REGION Network 25: RESET TEMPO DE OPERAÇÃO (HORAS)
   RUNG wire#powerrail
      Contact( #AUX09 )
      wire#w1
      { S7_GenerateENO := "TRUE" } Move(in := 0, out1 => #HOR)
   END_RUNG
   RUNG wire#powerrail
      Contact( #CRTO )
   END_RUNG wire#w1
   // the same network as SCL:
   IF #AUX09 OR #CRTO THEN #HOR := 0; END_IF;
END_REGION

REGION Network 26 (STL): ESCRITA DOS DADOS NO INVERSOR (PALAVRA DE COMANDO)
         A     "AlwaysTRUE";
         =     #CTW.DCbrakeRamp;
         =     #CTW.Coasting;
         =     #CTW.Enable_Ramp;
         =     #CTW.Enable_ramp_generator;
         =     #CTW.Control_plc;  //Valida setpoint


         A     #CL;
         =     #CTW.Start;  //LIGA/DESL

         A     #CL;
         A     #AUX10;
         A     #HAR;
         =     #CTW.Start_reverse;  //LIGA/DESL REVERSO


         A     #RESET;
         AN    #CL;
         =     #CTW.Reset;  //RESET
END_REGION
END_FUNCTION_BLOCK

FUNCTION_BLOCK "PDIR"   // FB207, LAD
{ S7_Optimized_Access := 'FALSE' }
VERSION : 0.1
   VAR_INPUT
      ML : Bool;
      MR : Bool;
      DL : Bool;
      MF1 : Bool;
      MF2 : Bool;
      HM : Bool;
      HA : Bool;
      CMA : Bool;
      CLM : Bool;
      CDM : Bool;
      CRF : Bool;
      CRTO : Bool;
      CL1S : Bool;
   END_VAR
   VAR_OUTPUT
      YFPP : Bool;
      YF : Bool;
      CL : Bool;
   END_VAR
   VAR_IN_OUT
      SEG : Int;
      MIN : Int;
      HOR : Int;
   END_VAR
   VAR
      AUX01 : Bool;
      AUX02 : Bool;
      AUX03 : Bool;
      AUX04 : Bool;
      AUX05 : Bool;
      AUX06 : Bool;
      AUX07 : Bool;
      AUX08 : Bool;
      AUX09 : Bool;
      P60S : Bool;
      P60M : Bool;
      PFHO : Bool;
      TPP1 : TON_TIME;
      TPP2 : TON_TIME;
   END_VAR
   VAR_TEMP
      TEMP0 : Bool;
      TEMP1 : Bool;
      ET_TPP1 : Time;
      ET_TPP2 : Time;
   END_VAR
   VAR_TEMP   // added for the SCL form of the ladder/FBD networks
      _w1 : Bool;
      _w2 : Bool;
      _w3 : Bool;
      _w4 : Bool;
   END_VAR
BEGIN

REGION Network 1: Falha na partida
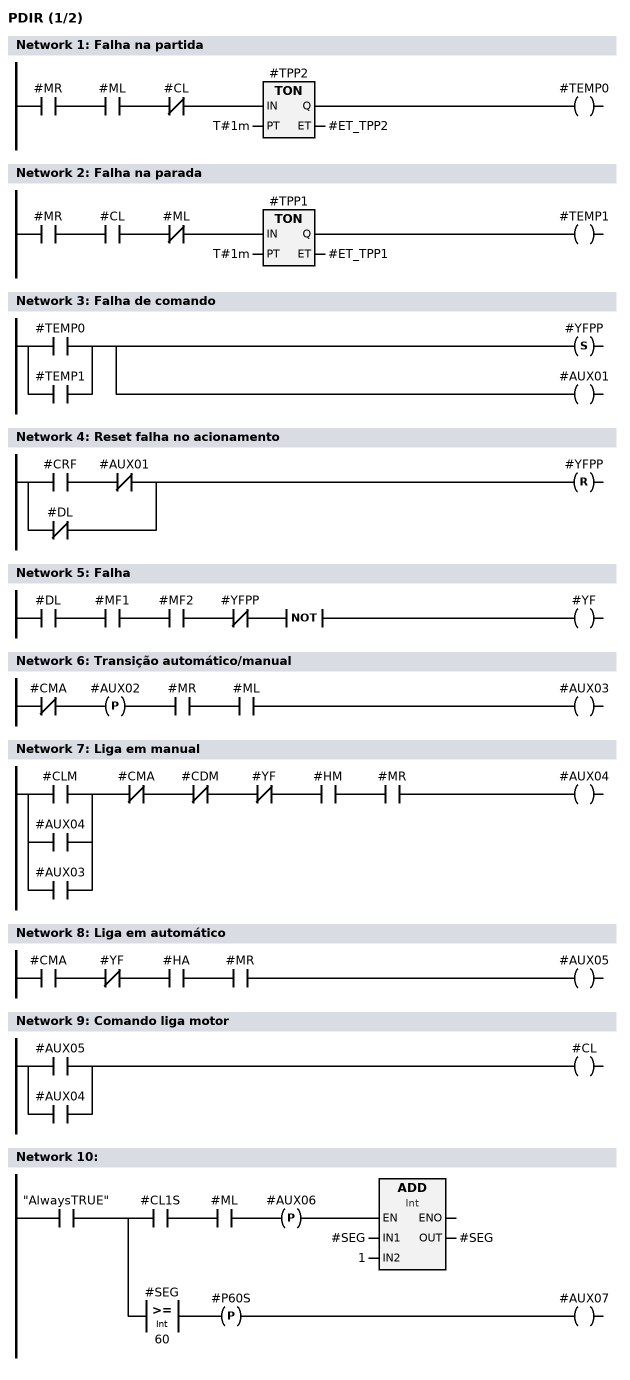
   #TPP2(IN := #MR AND #ML AND NOT #CL, PT := T#1m, ET => #ET_TPP2);   // TON
   #TEMP0 := #TPP2.Q;
END_REGION

REGION Network 2: Falha na parada
   #TPP1(IN := #MR AND #CL AND NOT #ML, PT := T#1m, ET => #ET_TPP1);   // TON
   #TEMP1 := #TPP1.Q;
END_REGION

REGION Network 3: Falha de comando
   RUNG wire#powerrail
      Contact( #TEMP0 )
      wire#w1
      S_Coil( #YFPP )
   END_RUNG
   RUNG wire#powerrail
      Contact( #TEMP1 )
   END_RUNG wire#w1
   RUNG wire#w1
      Coil( #AUX01 )
   END_RUNG
   // the same network as SCL:
   #_w1 := #TEMP0 OR #TEMP1;
   IF #_w1 THEN #YFPP := TRUE; END_IF;
   #AUX01 := #_w1;
END_REGION

REGION Network 4: Reset falha no acionamento
   RUNG wire#powerrail
      Contact( #CRF )
      I_Contact( #AUX01 )
      wire#w1
      R_Coil( #YFPP )
   END_RUNG
   RUNG wire#powerrail
      I_Contact( #DL )
   END_RUNG wire#w1
   // the same network as SCL:
   IF (#CRF AND NOT #AUX01) OR NOT #DL THEN #YFPP := FALSE; END_IF;
END_REGION

REGION Network 5: Falha
   RUNG wire#powerrail
      Contact( #DL )
      Contact( #MF1 )
      Contact( #MF2 )
      I_Contact( #YFPP )
      Not()
      Coil( #YF )
   END_RUNG
   // the same network as SCL:
   #YF := NOT (#DL AND #MF1 AND #MF2 AND NOT #YFPP);
END_REGION

REGION Network 6: Transição automático/manual
   RUNG wire#powerrail
      I_Contact( #CMA )
      P_Trig( #AUX02 )
      Contact( #MR )
      Contact( #ML )
      Coil( #AUX03 )
   END_RUNG
   // the same network as SCL:
   #_w1 := NOT #CMA AND NOT #AUX02;   // rising edge
   #AUX02 := NOT #CMA;
   #AUX03 := #_w1 AND #MR AND #ML;
END_REGION

REGION Network 7: Liga em manual
   RUNG wire#powerrail
      Contact( #CLM )
      wire#w1
      I_Contact( #CMA )
      I_Contact( #CDM )
      I_Contact( #YF )
      Contact( #HM )
      Contact( #MR )
      Coil( #AUX04 )
   END_RUNG
   RUNG wire#powerrail
      Contact( #AUX04 )
   END_RUNG wire#w1
   RUNG wire#powerrail
      Contact( #AUX03 )
   END_RUNG wire#w1
   // the same network as SCL:
   #AUX04 := (#CLM OR #AUX04 OR #AUX03) AND NOT #CMA AND NOT #CDM AND NOT #YF AND #HM AND #MR;
END_REGION

REGION Network 8: Liga em automático
   RUNG wire#powerrail
      Contact( #CMA )
      I_Contact( #YF )
      Contact( #HA )
      Contact( #MR )
      Coil( #AUX05 )
   END_RUNG
   // the same network as SCL:
   #AUX05 := #CMA AND NOT #YF AND #HA AND #MR;
END_REGION

REGION Network 9: Comando liga motor
   RUNG wire#powerrail
      Contact( #AUX05 )
      wire#w1
      Coil( #CL )
   END_RUNG
   RUNG wire#powerrail
      Contact( #AUX04 )
   END_RUNG wire#w1
   // the same network as SCL:
   #CL := #AUX05 OR #AUX04;
END_REGION

REGION Network 10
   RUNG wire#powerrail
      Contact( "AlwaysTRUE" )
      wire#w1
      Contact( #CL1S )
      Contact( #ML )
      P_Trig( #AUX06 )
      { S7_Templates := "SrcType := Int"; S7_GenerateENO := "TRUE" } Add(in1 := #SEG, in2 := 1, out => #SEG)
   END_RUNG
   RUNG wire#w1
      { S7_Templates := "SrcType := Int" } GE_Contact(in1 := #SEG, in2 := 60)
      P_Trig( #P60S )
      Coil( #AUX07 )
   END_RUNG
   // the same network as SCL:
   #_w1 := "AlwaysTRUE" AND #CL1S AND #ML;
   #_w2 := #_w1 AND NOT #AUX06;   // rising edge
   #AUX06 := #_w1;
   IF #_w2 THEN #SEG := #SEG + 1; END_IF;
   #_w3 := "AlwaysTRUE" AND (#SEG >= 60);
   #_w4 := #_w3 AND NOT #P60S;   // rising edge
   #P60S := #_w3;
   #AUX07 := #_w4;
END_REGION

REGION Network 11
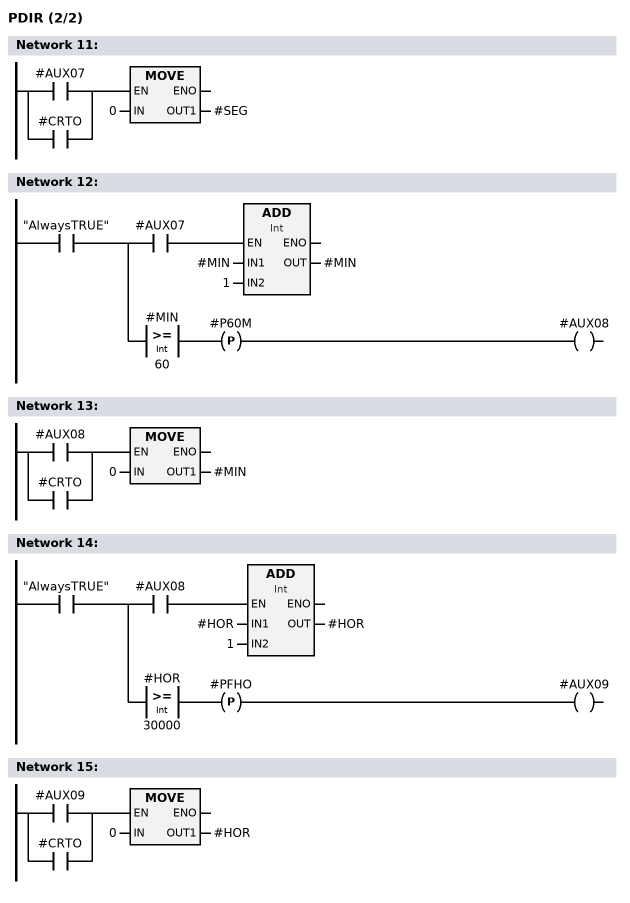
   RUNG wire#powerrail
      Contact( #AUX07 )
      wire#w1
      { S7_GenerateENO := "TRUE" } Move(in := 0, out1 => #SEG)
   END_RUNG
   RUNG wire#powerrail
      Contact( #CRTO )
   END_RUNG wire#w1
   // the same network as SCL:
   IF #AUX07 OR #CRTO THEN #SEG := 0; END_IF;
END_REGION

REGION Network 12
   RUNG wire#powerrail
      Contact( "AlwaysTRUE" )
      wire#w1
      Contact( #AUX07 )
      { S7_Templates := "SrcType := Int"; S7_GenerateENO := "TRUE" } Add(in1 := #MIN, in2 := 1, out => #MIN)
   END_RUNG
   RUNG wire#w1
      { S7_Templates := "SrcType := Int" } GE_Contact(in1 := #MIN, in2 := 60)
      P_Trig( #P60M )
      Coil( #AUX08 )
   END_RUNG
   // the same network as SCL:
   IF "AlwaysTRUE" AND #AUX07 THEN #MIN := #MIN + 1; END_IF;
   #_w1 := "AlwaysTRUE" AND (#MIN >= 60);
   #_w2 := #_w1 AND NOT #P60M;   // rising edge
   #P60M := #_w1;
   #AUX08 := #_w2;
END_REGION

REGION Network 13
   RUNG wire#powerrail
      Contact( #AUX08 )
      wire#w1
      { S7_GenerateENO := "TRUE" } Move(in := 0, out1 => #MIN)
   END_RUNG
   RUNG wire#powerrail
      Contact( #CRTO )
   END_RUNG wire#w1
   // the same network as SCL:
   IF #AUX08 OR #CRTO THEN #MIN := 0; END_IF;
END_REGION

REGION Network 14
   RUNG wire#powerrail
      Contact( "AlwaysTRUE" )
      wire#w1
      Contact( #AUX08 )
      { S7_Templates := "SrcType := Int"; S7_GenerateENO := "TRUE" } Add(in1 := #HOR, in2 := 1, out => #HOR)
   END_RUNG
   RUNG wire#w1
      { S7_Templates := "SrcType := Int" } GE_Contact(in1 := #HOR, in2 := 30000)
      P_Trig( #PFHO )
      Coil( #AUX09 )
   END_RUNG
   // the same network as SCL:
   IF "AlwaysTRUE" AND #AUX08 THEN #HOR := #HOR + 1; END_IF;
   #_w1 := "AlwaysTRUE" AND (#HOR >= 30000);
   #_w2 := #_w1 AND NOT #PFHO;   // rising edge
   #PFHO := #_w1;
   #AUX09 := #_w2;
END_REGION

REGION Network 15
   RUNG wire#powerrail
      Contact( #AUX09 )
      wire#w1
      { S7_GenerateENO := "TRUE" } Move(in := 0, out1 => #HOR)
   END_RUNG
   RUNG wire#powerrail
      Contact( #CRTO )
   END_RUNG wire#w1
   // the same network as SCL:
   IF #AUX09 OR #CRTO THEN #HOR := 0; END_IF;
END_REGION
END_FUNCTION_BLOCK

FUNCTION "IO" : Void   // FC1, LAD
{ S7_Optimized_Access := 'TRUE' }
VERSION : 0.1
BEGIN

REGION Network 1: Status e alarme elevatória principal 1
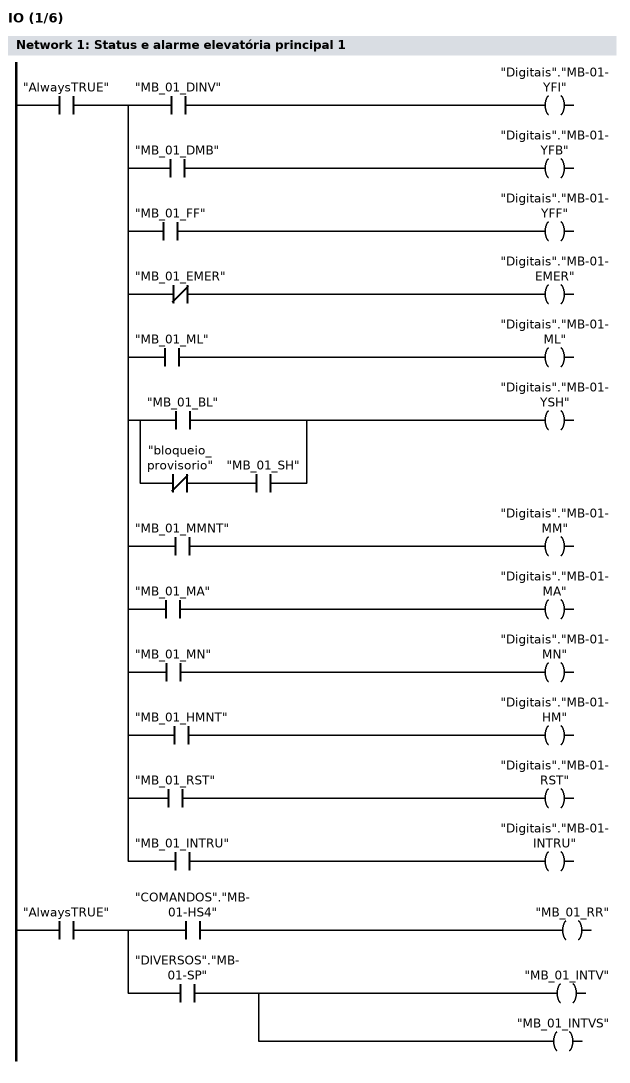
   RUNG wire#powerrail
      Contact( "AlwaysTRUE" )
      wire#w1
      Contact( "MB_01_DINV" )
      Coil( "Digitais"."MB-01-YFI" )
   END_RUNG
   RUNG wire#w1
      Contact( "MB_01_DMB" )
      Coil( "Digitais"."MB-01-YFB" )
   END_RUNG
   RUNG wire#w1
      Contact( "MB_01_FF" )
      Coil( "Digitais"."MB-01-YFF" )
   END_RUNG
   RUNG wire#w1
      I_Contact( "MB_01_EMER" )
      Coil( "Digitais"."MB-01-EMER" )
   END_RUNG
   RUNG wire#w1
      Contact( "MB_01_ML" )
      Coil( "Digitais"."MB-01-ML" )
   END_RUNG
   RUNG wire#w1
      Contact( "MB_01_BL" )
      wire#w2
      Coil( "Digitais"."MB-01-YSH" )
   END_RUNG
   RUNG wire#w1
      I_Contact( "bloqueio_provisorio" )
      Contact( "MB_01_SH" )
   END_RUNG wire#w2
   RUNG wire#w1
      Contact( "MB_01_MMNT" )
      Coil( "Digitais"."MB-01-MM" )
   END_RUNG
   RUNG wire#w1
      Contact( "MB_01_MA" )
      Coil( "Digitais"."MB-01-MA" )
   END_RUNG
   RUNG wire#w1
      Contact( "MB_01_MN" )
      Coil( "Digitais"."MB-01-MN" )
   END_RUNG
   RUNG wire#w1
      Contact( "MB_01_HMNT" )
      Coil( "Digitais"."MB-01-HM" )
   END_RUNG
   RUNG wire#w1
      Contact( "MB_01_RST" )
      Coil( "Digitais"."MB-01-RST" )
   END_RUNG
   RUNG wire#w1
      Contact( "MB_01_INTRU" )
      Coil( "Digitais"."MB-01-INTRU" )
   END_RUNG
   RUNG wire#powerrail
      Contact( "AlwaysTRUE" )
      wire#w3
      Contact( "COMANDOS"."MB-01-HS4" )
      Coil( "MB_01_RR" )
   END_RUNG
   RUNG wire#w3
      Contact( "DIVERSOS"."MB-01-SP" )
      wire#w4
      Coil( "MB_01_INTV" )
   END_RUNG
   RUNG wire#w4
      Coil( "MB_01_INTVS" )
   END_RUNG
   // the same network as SCL:
   "Digitais"."MB-01-YFI" := "AlwaysTRUE" AND "MB_01_DINV";
   "Digitais"."MB-01-YFB" := "AlwaysTRUE" AND "MB_01_DMB";
   "Digitais"."MB-01-YFF" := "AlwaysTRUE" AND "MB_01_FF";
   "Digitais"."MB-01-EMER" := "AlwaysTRUE" AND NOT "MB_01_EMER";
   "Digitais"."MB-01-ML" := "AlwaysTRUE" AND "MB_01_ML";
   "Digitais"."MB-01-YSH" := "AlwaysTRUE" AND ("MB_01_BL" OR (NOT "bloqueio_provisorio" AND "MB_01_SH"));
   "Digitais"."MB-01-MM" := "AlwaysTRUE" AND "MB_01_MMNT";
   "Digitais"."MB-01-MA" := "AlwaysTRUE" AND "MB_01_MA";
   "Digitais"."MB-01-MN" := "AlwaysTRUE" AND "MB_01_MN";
   "Digitais"."MB-01-HM" := "AlwaysTRUE" AND "MB_01_HMNT";
   "Digitais"."MB-01-RST" := "AlwaysTRUE" AND "MB_01_RST";
   "Digitais"."MB-01-INTRU" := "AlwaysTRUE" AND "MB_01_INTRU";
   "MB_01_RR" := "AlwaysTRUE" AND "COMANDOS"."MB-01-HS4";
   "MB_01_INTV" := "AlwaysTRUE" AND "DIVERSOS"."MB-01-SP";
   "MB_01_INTVS" := "MB_01_INTV";
END_REGION

REGION Network 2: Status e alarme elevatória principal 2
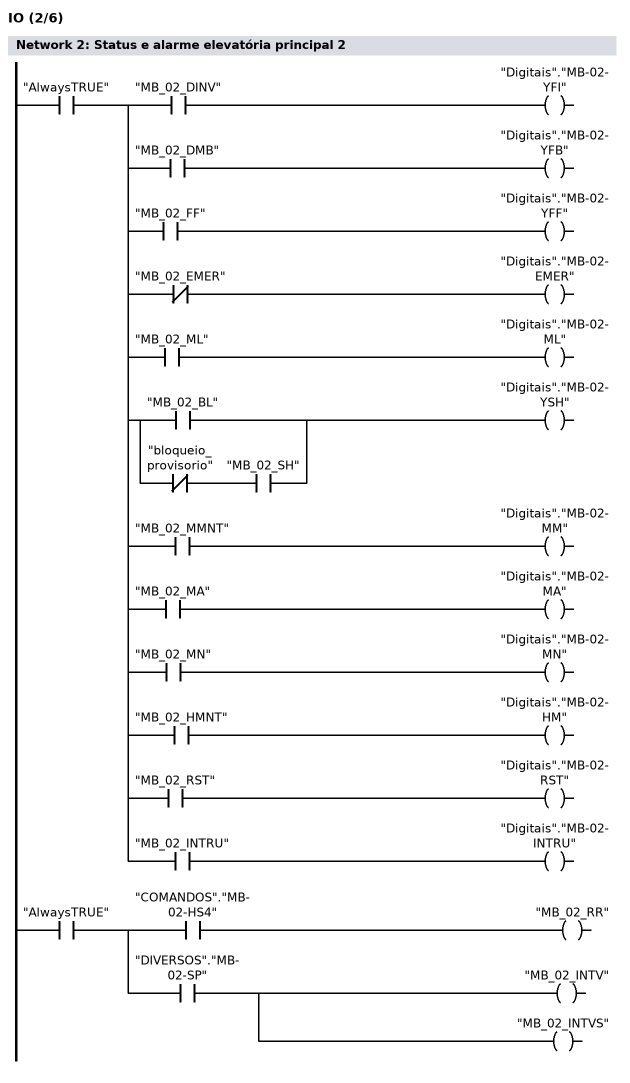
   RUNG wire#powerrail
      Contact( "AlwaysTRUE" )
      wire#w1
      Contact( "MB_02_DINV" )
      Coil( "Digitais"."MB-02-YFI" )
   END_RUNG
   RUNG wire#w1
      Contact( "MB_02_DMB" )
      Coil( "Digitais"."MB-02-YFB" )
   END_RUNG
   RUNG wire#w1
      Contact( "MB_02_FF" )
      Coil( "Digitais"."MB-02-YFF" )
   END_RUNG
   RUNG wire#w1
      I_Contact( "MB_02_EMER" )
      Coil( "Digitais"."MB-02-EMER" )
   END_RUNG
   RUNG wire#w1
      Contact( "MB_02_ML" )
      Coil( "Digitais"."MB-02-ML" )
   END_RUNG
   RUNG wire#w1
      Contact( "MB_02_BL" )
      wire#w2
      Coil( "Digitais"."MB-02-YSH" )
   END_RUNG
   RUNG wire#w1
      I_Contact( "bloqueio_provisorio" )
      Contact( "MB_02_SH" )
   END_RUNG wire#w2
   RUNG wire#w1
      Contact( "MB_02_MMNT" )
      Coil( "Digitais"."MB-02-MM" )
   END_RUNG
   RUNG wire#w1
      Contact( "MB_02_MA" )
      Coil( "Digitais"."MB-02-MA" )
   END_RUNG
   RUNG wire#w1
      Contact( "MB_02_MN" )
      Coil( "Digitais"."MB-02-MN" )
   END_RUNG
   RUNG wire#w1
      Contact( "MB_02_HMNT" )
      Coil( "Digitais"."MB-02-HM" )
   END_RUNG
   RUNG wire#w1
      Contact( "MB_02_RST" )
      Coil( "Digitais"."MB-02-RST" )
   END_RUNG
   RUNG wire#w1
      Contact( "MB_02_INTRU" )
      Coil( "Digitais"."MB-02-INTRU" )
   END_RUNG
   RUNG wire#powerrail
      Contact( "AlwaysTRUE" )
      wire#w3
      Contact( "COMANDOS"."MB-02-HS4" )
      Coil( "MB_02_RR" )
   END_RUNG
   RUNG wire#w3
      Contact( "DIVERSOS"."MB-02-SP" )
      wire#w4
      Coil( "MB_02_INTV" )
   END_RUNG
   RUNG wire#w4
      Coil( "MB_02_INTVS" )
   END_RUNG
   // the same network as SCL:
   "Digitais"."MB-02-YFI" := "AlwaysTRUE" AND "MB_02_DINV";
   "Digitais"."MB-02-YFB" := "AlwaysTRUE" AND "MB_02_DMB";
   "Digitais"."MB-02-YFF" := "AlwaysTRUE" AND "MB_02_FF";
   "Digitais"."MB-02-EMER" := "AlwaysTRUE" AND NOT "MB_02_EMER";
   "Digitais"."MB-02-ML" := "AlwaysTRUE" AND "MB_02_ML";
   "Digitais"."MB-02-YSH" := "AlwaysTRUE" AND ("MB_02_BL" OR (NOT "bloqueio_provisorio" AND "MB_02_SH"));
   "Digitais"."MB-02-MM" := "AlwaysTRUE" AND "MB_02_MMNT";
   "Digitais"."MB-02-MA" := "AlwaysTRUE" AND "MB_02_MA";
   "Digitais"."MB-02-MN" := "AlwaysTRUE" AND "MB_02_MN";
   "Digitais"."MB-02-HM" := "AlwaysTRUE" AND "MB_02_HMNT";
   "Digitais"."MB-02-RST" := "AlwaysTRUE" AND "MB_02_RST";
   "Digitais"."MB-02-INTRU" := "AlwaysTRUE" AND "MB_02_INTRU";
   "MB_02_RR" := "AlwaysTRUE" AND "COMANDOS"."MB-02-HS4";
   "MB_02_INTV" := "AlwaysTRUE" AND "DIVERSOS"."MB-02-SP";
   "MB_02_INTVS" := "MB_02_INTV";
END_REGION

REGION Network 3: Status e alarme elevatória principal 3
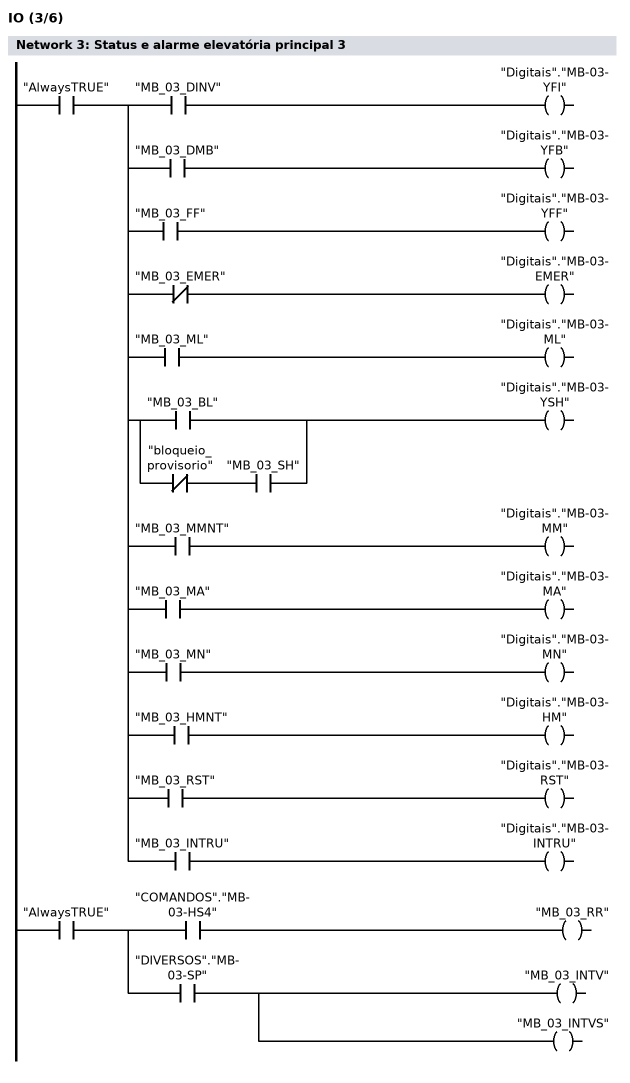
   RUNG wire#powerrail
      Contact( "AlwaysTRUE" )
      wire#w1
      Contact( "MB_03_DINV" )
      Coil( "Digitais"."MB-03-YFI" )
   END_RUNG
   RUNG wire#w1
      Contact( "MB_03_DMB" )
      Coil( "Digitais"."MB-03-YFB" )
   END_RUNG
   RUNG wire#w1
      Contact( "MB_03_FF" )
      Coil( "Digitais"."MB-03-YFF" )
   END_RUNG
   RUNG wire#w1
      I_Contact( "MB_03_EMER" )
      Coil( "Digitais"."MB-03-EMER" )
   END_RUNG
   RUNG wire#w1
      Contact( "MB_03_ML" )
      Coil( "Digitais"."MB-03-ML" )
   END_RUNG
   RUNG wire#w1
      Contact( "MB_03_BL" )
      wire#w2
      Coil( "Digitais"."MB-03-YSH" )
   END_RUNG
   RUNG wire#w1
      I_Contact( "bloqueio_provisorio" )
      Contact( "MB_03_SH" )
   END_RUNG wire#w2
   RUNG wire#w1
      Contact( "MB_03_MMNT" )
      Coil( "Digitais"."MB-03-MM" )
   END_RUNG
   RUNG wire#w1
      Contact( "MB_03_MA" )
      Coil( "Digitais"."MB-03-MA" )
   END_RUNG
   RUNG wire#w1
      Contact( "MB_03_MN" )
      Coil( "Digitais"."MB-03-MN" )
   END_RUNG
   RUNG wire#w1
      Contact( "MB_03_HMNT" )
      Coil( "Digitais"."MB-03-HM" )
   END_RUNG
   RUNG wire#w1
      Contact( "MB_03_RST" )
      Coil( "Digitais"."MB-03-RST" )
   END_RUNG
   RUNG wire#w1
      Contact( "MB_03_INTRU" )
      Coil( "Digitais"."MB-03-INTRU" )
   END_RUNG
   RUNG wire#powerrail
      Contact( "AlwaysTRUE" )
      wire#w3
      Contact( "COMANDOS"."MB-03-HS4" )
      Coil( "MB_03_RR" )
   END_RUNG
   RUNG wire#w3
      Contact( "DIVERSOS"."MB-03-SP" )
      wire#w4
      Coil( "MB_03_INTV" )
   END_RUNG
   RUNG wire#w4
      Coil( "MB_03_INTVS" )
   END_RUNG
   // the same network as SCL:
   "Digitais"."MB-03-YFI" := "AlwaysTRUE" AND "MB_03_DINV";
   "Digitais"."MB-03-YFB" := "AlwaysTRUE" AND "MB_03_DMB";
   "Digitais"."MB-03-YFF" := "AlwaysTRUE" AND "MB_03_FF";
   "Digitais"."MB-03-EMER" := "AlwaysTRUE" AND NOT "MB_03_EMER";
   "Digitais"."MB-03-ML" := "AlwaysTRUE" AND "MB_03_ML";
   "Digitais"."MB-03-YSH" := "AlwaysTRUE" AND ("MB_03_BL" OR (NOT "bloqueio_provisorio" AND "MB_03_SH"));
   "Digitais"."MB-03-MM" := "AlwaysTRUE" AND "MB_03_MMNT";
   "Digitais"."MB-03-MA" := "AlwaysTRUE" AND "MB_03_MA";
   "Digitais"."MB-03-MN" := "AlwaysTRUE" AND "MB_03_MN";
   "Digitais"."MB-03-HM" := "AlwaysTRUE" AND "MB_03_HMNT";
   "Digitais"."MB-03-RST" := "AlwaysTRUE" AND "MB_03_RST";
   "Digitais"."MB-03-INTRU" := "AlwaysTRUE" AND "MB_03_INTRU";
   "MB_03_RR" := "AlwaysTRUE" AND "COMANDOS"."MB-03-HS4";
   "MB_03_INTV" := "AlwaysTRUE" AND "DIVERSOS"."MB-03-SP";
   "MB_03_INTVS" := "MB_03_INTV";
END_REGION

REGION Network 4: Status e alarme elevatória principal 4
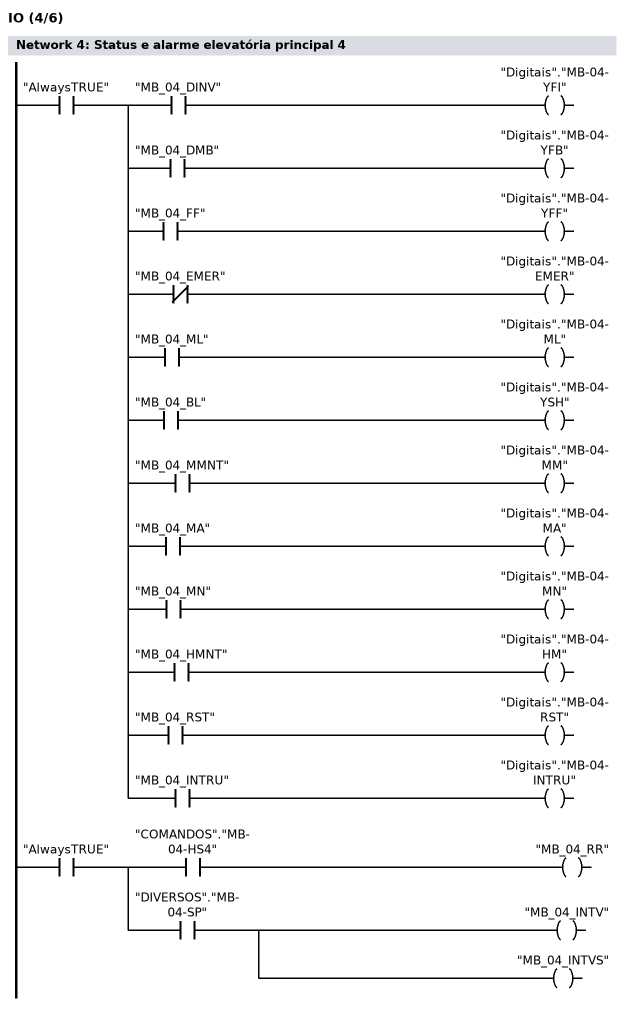
   RUNG wire#powerrail
      Contact( "AlwaysTRUE" )
      wire#w1
      Contact( "MB_04_DINV" )
      Coil( "Digitais"."MB-04-YFI" )
   END_RUNG
   RUNG wire#w1
      Contact( "MB_04_DMB" )
      Coil( "Digitais"."MB-04-YFB" )
   END_RUNG
   RUNG wire#w1
      Contact( "MB_04_FF" )
      Coil( "Digitais"."MB-04-YFF" )
   END_RUNG
   RUNG wire#w1
      I_Contact( "MB_04_EMER" )
      Coil( "Digitais"."MB-04-EMER" )
   END_RUNG
   RUNG wire#w1
      Contact( "MB_04_ML" )
      Coil( "Digitais"."MB-04-ML" )
   END_RUNG
   RUNG wire#w1
      Contact( "MB_04_BL" )
      Coil( "Digitais"."MB-04-YSH" )
   END_RUNG
   RUNG wire#w1
      Contact( "MB_04_MMNT" )
      Coil( "Digitais"."MB-04-MM" )
   END_RUNG
   RUNG wire#w1
      Contact( "MB_04_MA" )
      Coil( "Digitais"."MB-04-MA" )
   END_RUNG
   RUNG wire#w1
      Contact( "MB_04_MN" )
      Coil( "Digitais"."MB-04-MN" )
   END_RUNG
   RUNG wire#w1
      Contact( "MB_04_HMNT" )
      Coil( "Digitais"."MB-04-HM" )
   END_RUNG
   RUNG wire#w1
      Contact( "MB_04_RST" )
      Coil( "Digitais"."MB-04-RST" )
   END_RUNG
   RUNG wire#w1
      Contact( "MB_04_INTRU" )
      Coil( "Digitais"."MB-04-INTRU" )
   END_RUNG
   RUNG wire#powerrail
      Contact( "AlwaysTRUE" )
      wire#w2
      Contact( "COMANDOS"."MB-04-HS4" )
      Coil( "MB_04_RR" )
   END_RUNG
   RUNG wire#w2
      Contact( "DIVERSOS"."MB-04-SP" )
      wire#w3
      Coil( "MB_04_INTV" )
   END_RUNG
   RUNG wire#w3
      Coil( "MB_04_INTVS" )
   END_RUNG
   // the same network as SCL:
   "Digitais"."MB-04-YFI" := "AlwaysTRUE" AND "MB_04_DINV";
   "Digitais"."MB-04-YFB" := "AlwaysTRUE" AND "MB_04_DMB";
   "Digitais"."MB-04-YFF" := "AlwaysTRUE" AND "MB_04_FF";
   "Digitais"."MB-04-EMER" := "AlwaysTRUE" AND NOT "MB_04_EMER";
   "Digitais"."MB-04-ML" := "AlwaysTRUE" AND "MB_04_ML";
   "Digitais"."MB-04-YSH" := "AlwaysTRUE" AND "MB_04_BL";
   "Digitais"."MB-04-MM" := "AlwaysTRUE" AND "MB_04_MMNT";
   "Digitais"."MB-04-MA" := "AlwaysTRUE" AND "MB_04_MA";
   "Digitais"."MB-04-MN" := "AlwaysTRUE" AND "MB_04_MN";
   "Digitais"."MB-04-HM" := "AlwaysTRUE" AND "MB_04_HMNT";
   "Digitais"."MB-04-RST" := "AlwaysTRUE" AND "MB_04_RST";
   "Digitais"."MB-04-INTRU" := "AlwaysTRUE" AND "MB_04_INTRU";
   "MB_04_RR" := "AlwaysTRUE" AND "COMANDOS"."MB-04-HS4";
   "MB_04_INTV" := "AlwaysTRUE" AND "DIVERSOS"."MB-04-SP";
   "MB_04_INTVS" := "MB_04_INTV";
END_REGION

REGION Network 5: Status e alarme PCM-E-CF-01-04
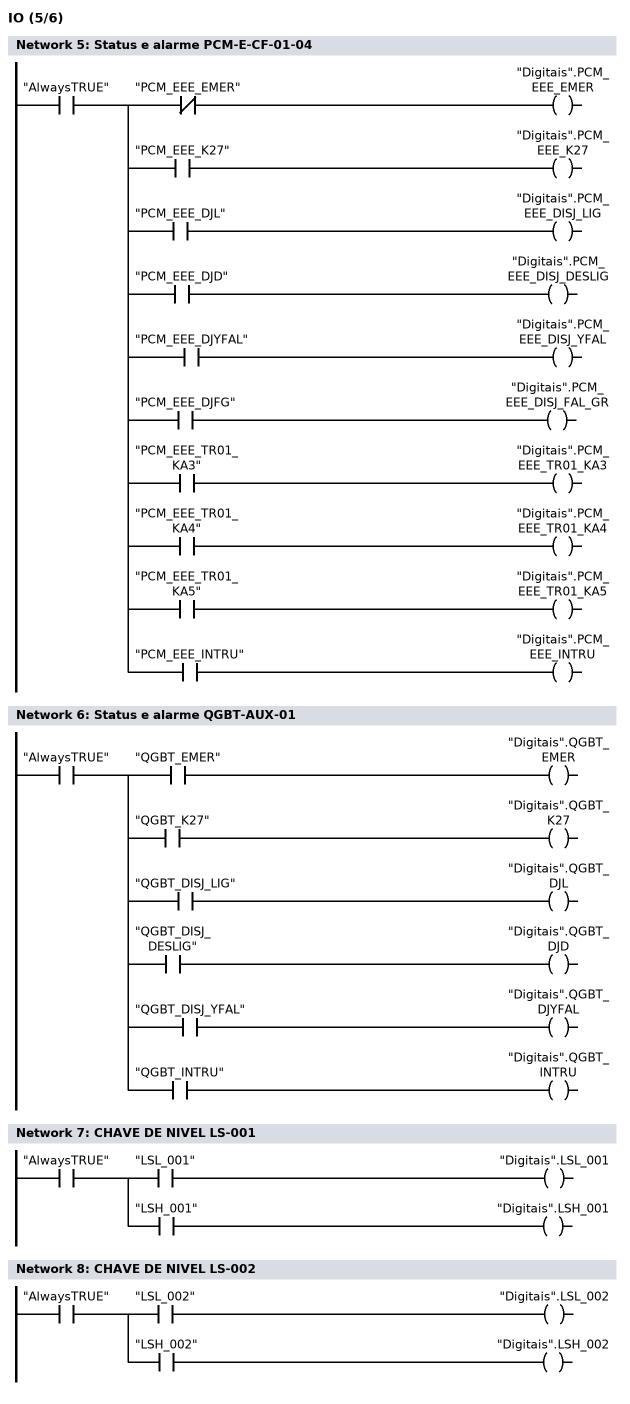
   RUNG wire#powerrail
      Contact( "AlwaysTRUE" )
      wire#w1
      I_Contact( "PCM_EEE_EMER" )
      Coil( "Digitais".PCM_EEE_EMER )
   END_RUNG
   RUNG wire#w1
      Contact( "PCM_EEE_K27" )
      Coil( "Digitais".PCM_EEE_K27 )
   END_RUNG
   RUNG wire#w1
      Contact( "PCM_EEE_DJL" )
      Coil( "Digitais".PCM_EEE_DISJ_LIG )
   END_RUNG
   RUNG wire#w1
      Contact( "PCM_EEE_DJD" )
      Coil( "Digitais".PCM_EEE_DISJ_DESLIG )
   END_RUNG
   RUNG wire#w1
      Contact( "PCM_EEE_DJYFAL" )
      Coil( "Digitais".PCM_EEE_DISJ_YFAL )
   END_RUNG
   RUNG wire#w1
      Contact( "PCM_EEE_DJFG" )
      Coil( "Digitais".PCM_EEE_DISJ_FAL_GR )
   END_RUNG
   RUNG wire#w1
      Contact( "PCM_EEE_TR01_KA3" )
      Coil( "Digitais".PCM_EEE_TR01_KA3 )
   END_RUNG
   RUNG wire#w1
      Contact( "PCM_EEE_TR01_KA4" )
      Coil( "Digitais".PCM_EEE_TR01_KA4 )
   END_RUNG
   RUNG wire#w1
      Contact( "PCM_EEE_TR01_KA5" )
      Coil( "Digitais".PCM_EEE_TR01_KA5 )
   END_RUNG
   RUNG wire#w1
      Contact( "PCM_EEE_INTRU" )
      Coil( "Digitais".PCM_EEE_INTRU )
   END_RUNG
   // the same network as SCL:
   "Digitais".PCM_EEE_EMER := "AlwaysTRUE" AND NOT "PCM_EEE_EMER";
   "Digitais".PCM_EEE_K27 := "AlwaysTRUE" AND "PCM_EEE_K27";
   "Digitais".PCM_EEE_DISJ_LIG := "AlwaysTRUE" AND "PCM_EEE_DJL";
   "Digitais".PCM_EEE_DISJ_DESLIG := "AlwaysTRUE" AND "PCM_EEE_DJD";
   "Digitais".PCM_EEE_DISJ_YFAL := "AlwaysTRUE" AND "PCM_EEE_DJYFAL";
   "Digitais".PCM_EEE_DISJ_FAL_GR := "AlwaysTRUE" AND "PCM_EEE_DJFG";
   "Digitais".PCM_EEE_TR01_KA3 := "AlwaysTRUE" AND "PCM_EEE_TR01_KA3";
   "Digitais".PCM_EEE_TR01_KA4 := "AlwaysTRUE" AND "PCM_EEE_TR01_KA4";
   "Digitais".PCM_EEE_TR01_KA5 := "AlwaysTRUE" AND "PCM_EEE_TR01_KA5";
   "Digitais".PCM_EEE_INTRU := "AlwaysTRUE" AND "PCM_EEE_INTRU";
END_REGION

REGION Network 6: Status e alarme QGBT-AUX-01
   RUNG wire#powerrail
      Contact( "AlwaysTRUE" )
      wire#w1
      Contact( "QGBT_EMER" )
      Coil( "Digitais".QGBT_EMER )
   END_RUNG
   RUNG wire#w1
      Contact( "QGBT_K27" )
      Coil( "Digitais".QGBT_K27 )
   END_RUNG
   RUNG wire#w1
      Contact( "QGBT_DISJ_LIG" )
      Coil( "Digitais".QGBT_DJL )
   END_RUNG
   RUNG wire#w1
      Contact( "QGBT_DISJ_DESLIG" )
      Coil( "Digitais".QGBT_DJD )
   END_RUNG
   RUNG wire#w1
      Contact( "QGBT_DISJ_YFAL" )
      Coil( "Digitais".QGBT_DJYFAL )
   END_RUNG
   RUNG wire#w1
      Contact( "QGBT_INTRU" )
      Coil( "Digitais".QGBT_INTRU )
   END_RUNG
   // the same network as SCL:
   "Digitais".QGBT_EMER := "AlwaysTRUE" AND "QGBT_EMER";
   "Digitais".QGBT_K27 := "AlwaysTRUE" AND "QGBT_K27";
   "Digitais".QGBT_DJL := "AlwaysTRUE" AND "QGBT_DISJ_LIG";
   "Digitais".QGBT_DJD := "AlwaysTRUE" AND "QGBT_DISJ_DESLIG";
   "Digitais".QGBT_DJYFAL := "AlwaysTRUE" AND "QGBT_DISJ_YFAL";
   "Digitais".QGBT_INTRU := "AlwaysTRUE" AND "QGBT_INTRU";
END_REGION

REGION Network 7: CHAVE DE NIVEL LS-001
   RUNG wire#powerrail
      Contact( "AlwaysTRUE" )
      wire#w1
      Contact( "LSL_001" )
      Coil( "Digitais".LSL_001 )
   END_RUNG
   RUNG wire#w1
      Contact( "LSH_001" )
      Coil( "Digitais".LSH_001 )
   END_RUNG
   // the same network as SCL:
   "Digitais".LSL_001 := "AlwaysTRUE" AND "LSL_001";
   "Digitais".LSH_001 := "AlwaysTRUE" AND "LSH_001";
END_REGION

REGION Network 8: CHAVE DE NIVEL LS-002
   RUNG wire#powerrail
      Contact( "AlwaysTRUE" )
      wire#w1
      Contact( "LSL_002" )
      Coil( "Digitais".LSL_002 )
   END_RUNG
   RUNG wire#w1
      Contact( "LSH_002" )
      Coil( "Digitais".LSH_002 )
   END_RUNG
   // the same network as SCL:
   "Digitais".LSL_002 := "AlwaysTRUE" AND "LSL_002";
   "Digitais".LSH_002 := "AlwaysTRUE" AND "LSH_002";
END_REGION

REGION Network 9: Status e alarme PCE-EEE
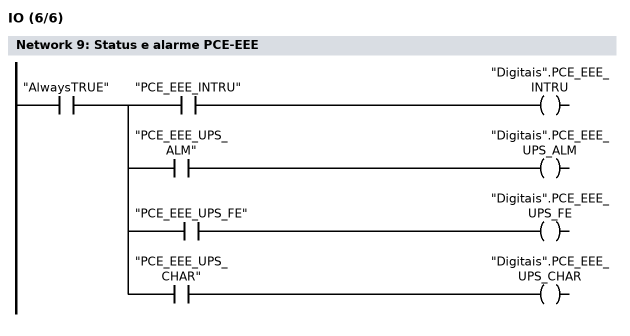
   RUNG wire#powerrail
      Contact( "AlwaysTRUE" )
      wire#w1
      Contact( "PCE_EEE_INTRU" )
      Coil( "Digitais".PCE_EEE_INTRU )
   END_RUNG
   RUNG wire#w1
      Contact( "PCE_EEE_UPS_ALM" )
      Coil( "Digitais".PCE_EEE_UPS_ALM )
   END_RUNG
   RUNG wire#w1
      Contact( "PCE_EEE_UPS_FE" )
      Coil( "Digitais".PCE_EEE_UPS_FE )
   END_RUNG
   RUNG wire#w1
      Contact( "PCE_EEE_UPS_CHAR" )
      Coil( "Digitais".PCE_EEE_UPS_CHAR )
   END_RUNG
   // the same network as SCL:
   "Digitais".PCE_EEE_INTRU := "AlwaysTRUE" AND "PCE_EEE_INTRU";
   "Digitais".PCE_EEE_UPS_ALM := "AlwaysTRUE" AND "PCE_EEE_UPS_ALM";
   "Digitais".PCE_EEE_UPS_FE := "AlwaysTRUE" AND "PCE_EEE_UPS_FE";
   "Digitais".PCE_EEE_UPS_CHAR := "AlwaysTRUE" AND "PCE_EEE_UPS_CHAR";
END_REGION
END_FUNCTION

FUNCTION "AlARME" : Void   // FC3, LAD
{ S7_Optimized_Access := 'TRUE' }
VERSION : 0.1
BEGIN

REGION Network 1: ALARMES IHM
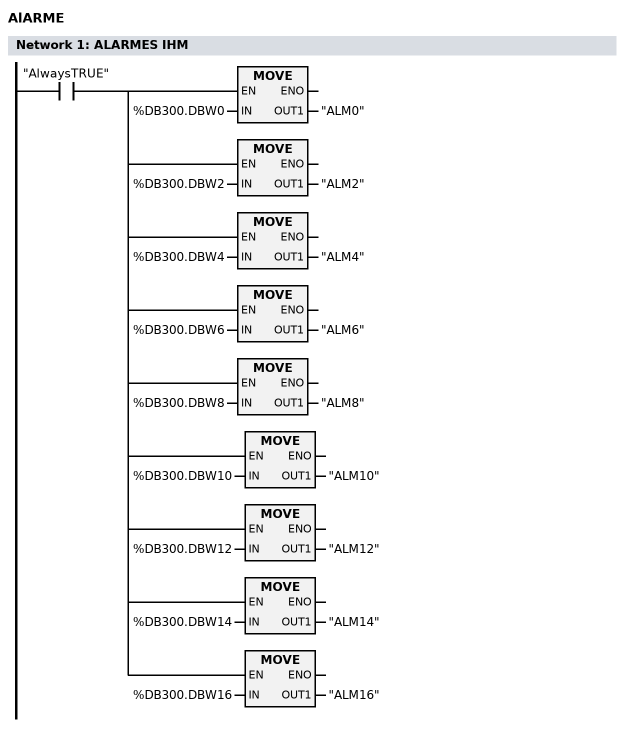
   RUNG wire#powerrail
      Contact( "AlwaysTRUE" )
      wire#w1
      Move(in := %DB300.DBW0, out1 => "ALM0")
   END_RUNG
   RUNG wire#w1
      Move(in := %DB300.DBW2, out1 => "ALM2")
   END_RUNG
   RUNG wire#w1
      Move(in := %DB300.DBW4, out1 => "ALM4")
   END_RUNG
   RUNG wire#w1
      Move(in := %DB300.DBW6, out1 => "ALM6")
   END_RUNG
   RUNG wire#w1
      Move(in := %DB300.DBW8, out1 => "ALM8")
   END_RUNG
   RUNG wire#w1
      Move(in := %DB300.DBW10, out1 => "ALM10")
   END_RUNG
   RUNG wire#w1
      Move(in := %DB300.DBW12, out1 => "ALM12")
   END_RUNG
   RUNG wire#w1
      Move(in := %DB300.DBW14, out1 => "ALM14")
   END_RUNG
   RUNG wire#w1
      Move(in := %DB300.DBW16, out1 => "ALM16")
   END_RUNG
   // the same network as SCL:
   IF "AlwaysTRUE" THEN
       "ALM0" := %DB300.DBW0;
       "ALM2" := %DB300.DBW2;
       "ALM4" := %DB300.DBW4;
       "ALM6" := %DB300.DBW6;
       "ALM8" := %DB300.DBW8;
       "ALM10" := %DB300.DBW10;
       "ALM12" := %DB300.DBW12;
       "ALM14" := %DB300.DBW14;
       "ALM16" := %DB300.DBW16;
   END_IF;
END_REGION
END_FUNCTION

FUNCTION "MB-01" : Void   // FC22, LAD
TITLE = Lógica de acionamento do motor
{ S7_Optimized_Access := 'FALSE' }
VERSION : 0.1
   VAR_TEMP
      IM : Bool;   // Intertravamento manual = 0
      IA : Bool;   // Intertravamento automáticol = 0
      HABM : Bool;   // Habilita funcionamento manual = 1
      HABA : Bool;   // Habilita funcionamento automático = 1
      CLM : Bool;   // Comando liga motor
      PROT : Bool;   // Proteção do motor acionada
   END_VAR
BEGIN

REGION Network 1: Intertravamento maual/automático
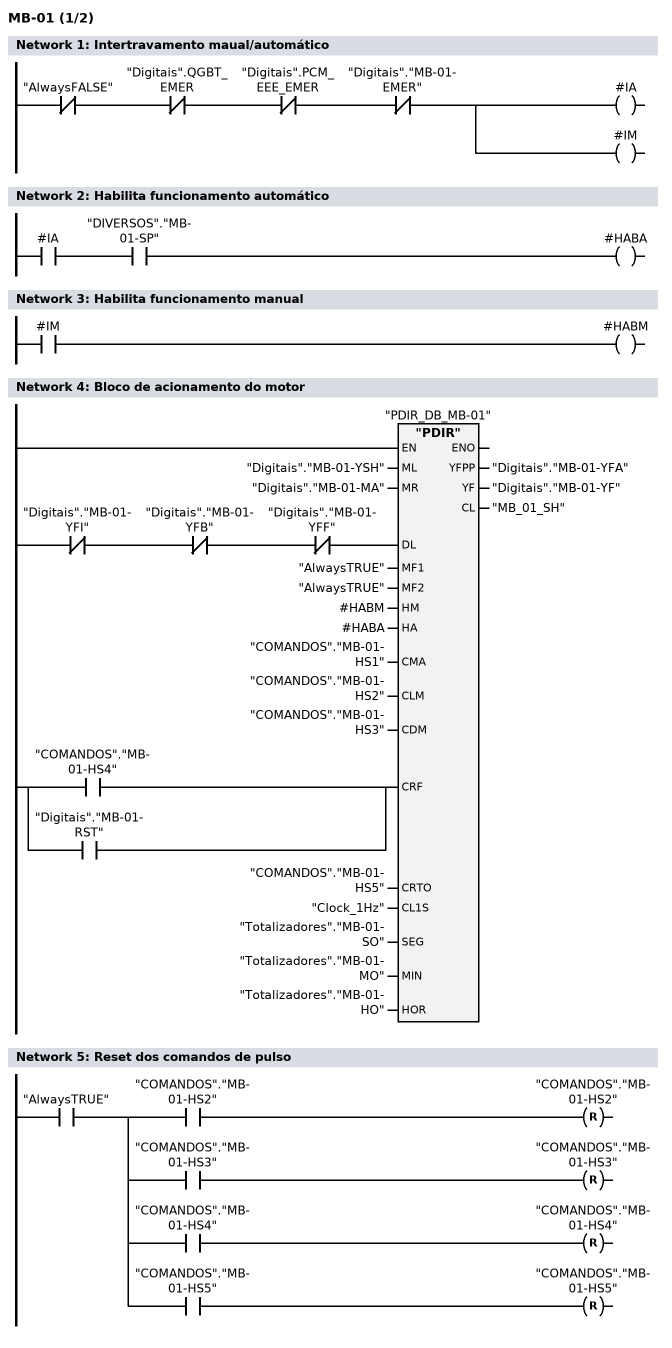
   RUNG wire#powerrail
      I_Contact( "AlwaysFALSE" )
      I_Contact( "Digitais".QGBT_EMER )
      I_Contact( "Digitais".PCM_EEE_EMER )
      I_Contact( "Digitais"."MB-01-EMER" )
      wire#w1
      Coil( #IA )
   END_RUNG
   RUNG wire#w1
      Coil( #IM )
   END_RUNG
   // the same network as SCL:
   #IA := NOT "AlwaysFALSE" AND NOT "Digitais".QGBT_EMER AND NOT "Digitais".PCM_EEE_EMER AND NOT "Digitais"."MB-01-EMER";
   #IM := #IA;
END_REGION

REGION Network 2: Habilita funcionamento automático
   RUNG wire#powerrail
      Contact( #IA )
      Contact( "DIVERSOS"."MB-01-SP" )
      Coil( #HABA )
   END_RUNG
   // the same network as SCL:
   #HABA := #IA AND "DIVERSOS"."MB-01-SP";
END_REGION

REGION Network 3: Habilita funcionamento manual
   RUNG wire#powerrail
      Contact( #IM )
      Coil( #HABM )
   END_RUNG
   // the same network as SCL:
   #HABM := #IM;
END_REGION

REGION Network 4: Bloco de acionamento do motor
   RUNG wire#powerrail
      "PDIR_DB_MB-01"(DL := wire#w1, CRF := wire#w2, ML := "Digitais"."MB-01-YSH", MR := "Digitais"."MB-01-MA", MF1 := "AlwaysTRUE", MF2 := "AlwaysTRUE", HM := #HABM, HA := #HABA, CMA := "COMANDOS"."MB-01-HS1", CLM := "COMANDOS"."MB-01-HS2", CDM := "COMANDOS"."MB-01-HS3", CRTO := "COMANDOS"."MB-01-HS5", CL1S := "Clock_1Hz", SEG := "Totalizadores"."MB-01-SO", MIN := "Totalizadores"."MB-01-MO", HOR := "Totalizadores"."MB-01-HO", YFPP => "Digitais"."MB-01-YFA", YF => "Digitais"."MB-01-YF", CL => "MB_01_SH")
   END_RUNG
   RUNG wire#powerrail
      I_Contact( "Digitais"."MB-01-YFI" )
      I_Contact( "Digitais"."MB-01-YFB" )
      I_Contact( "Digitais"."MB-01-YFF" )
   END_RUNG wire#w1
   RUNG wire#powerrail
      Contact( "COMANDOS"."MB-01-HS4" )
   END_RUNG wire#w2
   RUNG wire#powerrail
      Contact( "Digitais"."MB-01-RST" )
   END_RUNG wire#w2
   // the same network as SCL:
   "PDIR_DB_MB-01"(ML := "Digitais"."MB-01-YSH",   // "PDIR"
                   MR := "Digitais"."MB-01-MA",
                   DL := NOT "Digitais"."MB-01-YFI" AND NOT "Digitais"."MB-01-YFB" AND NOT "Digitais"."MB-01-YFF",
                   MF1 := "AlwaysTRUE",
                   MF2 := "AlwaysTRUE",
                   HM := #HABM,
                   HA := #HABA,
                   CMA := "COMANDOS"."MB-01-HS1",
                   CLM := "COMANDOS"."MB-01-HS2",
                   CDM := "COMANDOS"."MB-01-HS3",
                   CRF := "COMANDOS"."MB-01-HS4" OR "Digitais"."MB-01-RST",
                   CRTO := "COMANDOS"."MB-01-HS5",
                   CL1S := "Clock_1Hz",
                   SEG := "Totalizadores"."MB-01-SO",
                   MIN := "Totalizadores"."MB-01-MO",
                   HOR := "Totalizadores"."MB-01-HO",
                   YFPP => "Digitais"."MB-01-YFA",
                   YF => "Digitais"."MB-01-YF",
                   CL => "MB_01_SH");
END_REGION

REGION Network 5: Reset dos comandos de pulso
   RUNG wire#powerrail
      Contact( "AlwaysTRUE" )
      wire#w1
      Contact( "COMANDOS"."MB-01-HS2" )
      R_Coil( "COMANDOS"."MB-01-HS2" )
   END_RUNG
   RUNG wire#w1
      Contact( "COMANDOS"."MB-01-HS3" )
      R_Coil( "COMANDOS"."MB-01-HS3" )
   END_RUNG
   RUNG wire#w1
      Contact( "COMANDOS"."MB-01-HS4" )
      R_Coil( "COMANDOS"."MB-01-HS4" )
   END_RUNG
   RUNG wire#w1
      Contact( "COMANDOS"."MB-01-HS5" )
      R_Coil( "COMANDOS"."MB-01-HS5" )
   END_RUNG
   // the same network as SCL:
   IF "AlwaysTRUE" AND "COMANDOS"."MB-01-HS2" THEN "COMANDOS"."MB-01-HS2" := FALSE; END_IF;
   IF "AlwaysTRUE" AND "COMANDOS"."MB-01-HS3" THEN "COMANDOS"."MB-01-HS3" := FALSE; END_IF;
   IF "AlwaysTRUE" AND "COMANDOS"."MB-01-HS4" THEN "COMANDOS"."MB-01-HS4" := FALSE; END_IF;
   IF "AlwaysTRUE" AND "COMANDOS"."MB-01-HS5" THEN "COMANDOS"."MB-01-HS5" := FALSE; END_IF;
END_REGION

REGION Network 6: Elevatoria principal modo automatico
